FUNCTION_BLOCK "Sim: from Global"   // FB26, SCL
{ S7_Optimized_Access := 'TRUE' }
VERSION : 0.1
   VAR_INPUT
      stns : "Station: All Stations";
   END_VAR
   VAR_IN_OUT
      simStations : "Simulated Stations";
   END_VAR
   VAR
      old : Struct
         nextGrp : Bool;
         prevGrp : Bool;
      END_STRUCT;
   END_VAR
   VAR_TEMP
      animate : USInt;
      btnCount : Int;
      currentBtn : Bool;
      dzLabel : WString;
      firstStn : Int;
      i : Int;
      intBox : Int;
      j : Int;
      kp8Color : DWord;
      label : WString;
      oldBtn : Bool;
      pSim : Int;
      pStn : Int;
   END_VAR
   VAR CONSTANT
      space : WString := WSTRING#' ';
      lead0 : WString := WSTRING#'0';
      volvo16 : WString := WSTRING#'VOLVO 16';
   END_VAR
BEGIN
   REGION "COPY TO LOCAL"
       #firstStn := #simStations.firstStn;
   END_REGION

   REGION "RESOLVE STATION POINTER"

       REGION "PROCESS NEXT GROUP PRESS"

           REGION "COPY TO LOCAL"
               #currentBtn := #simStations.down.actuate;
               #oldBtn := #old.nextGrp;
           END_REGION

           REGION "FALLING EDGE OF NEXT GROUP"
               IF NOT #currentBtn AND #oldBtn THEN

                   REGION "INCREMENT FIRST STATION"
                       #firstStn += "simKP8Count";
                   END_REGION

                   REGION "UPPER LIMIT ROLL OVER"
                       IF #firstStn > "STATION_COUNT" THEN
                           #firstStn -= "STATION_COUNT" + 1;
                       END_IF;
                   END_REGION

               END_IF;
           END_REGION

           REGION "NEXT GROUP CHANGE DETECTION"
               #old.nextGrp := #currentBtn;
           END_REGION

       END_REGION

       REGION "PROCESS PREVIOUS GROUP PRESS"

           REGION "COPY TO LOCAL"
               #currentBtn := #simStations.up.actuate;
               #oldBtn := #old.prevGrp;
           END_REGION

           REGION "FALLING EDGE OF PREVIOUS GROUP"
               IF NOT #currentBtn AND #oldBtn THEN

                   REGION "DECREMENT FIRST STATION"
                       #firstStn -= "simKP8Count";
                   END_REGION

                   REGION "LOWER LIMIT ROLL OVER"
                       IF #firstStn < 0 THEN
                           #firstStn += "STATION_COUNT" + 1;
                       END_IF;
                   END_REGION

               END_IF;
           END_REGION

           REGION "PREVIOUS GROUP CHANGE DETECTION"
               #old.prevGrp := #currentBtn;
           END_REGION

       END_REGION

   END_REGION

   REGION "FOR EACH BUTTON"
       FOR #i := 0 TO 11 DO

           REGION "CALCULATE POINTER"
               #pStn := #i + #firstStn;
               #pSim := #i;
           END_REGION

           REGION "UPPER LIMIT ROLL OVER"
               IF #pStn > "STATION_COUNT" THEN
                   #pStn := #firstStn + #i - "STATION_COUNT" - 1;
               END_IF;
           END_REGION

           REGION "COPY TO LOCAL"
               #kp8Color := #stns.stn[#pStn].wipCmpts.ioData.kp8.tempOut;
           END_REGION

           REGION "LABEL STATIONS"

               REGION "DETERMINE LINE LABEL"
                   #label := #stns.stn[#pStn].id.lineName;
                   IF #label = #volvo16 THEN
                       #label := WSTRING#'V16';
                   END_IF;
               END_REGION

               REGION "DETERMINE DROP ZONE LABEL"
                   #intBox := USINT_TO_INT(#stns.stn[#pStn].id.dropZone);
                   IF #intBox <= 9 THEN
                       #dzLabel := CONCAT_WSTRING(IN1 := #lead0,
                                                  IN2 := "Strip Sign"(INT_TO_WSTRING(#intBox)));
                   END_IF;
                   IF #intBox >= 10 THEN
                       #dzLabel := "Strip Sign"(INT_TO_WSTRING(#intBox));
                   END_IF;
               END_REGION

               REGION "WRITE LABEL"
                   #label := CONCAT_WSTRING(IN1 := #label,
                                            IN2 := #space,
                                            IN3 := #dzLabel);
                   #simStations.me[#pSim].stn.label := #label;
               END_REGION

           END_REGION

           REGION "ANIMATE STATION LABEL"
               #simStations.me[#pSim].stn.animate := "GRAY_BACKGROUND";
           END_REGION

           REGION "FOR EACH BUTTON"
               FOR #j := 0 TO "BUTTON_COUNT" DO

                   REGION "COLOR BUTTONS"
                       #animate := "KP8 Driver: HMI Emulator: Animation"(kp8Color := #kp8Color,
                                                                btnNumber := #j);
                       #simStations.me[#pSim].btn.animate[#j] := #animate;
                   END_REGION

                   REGION "WRITE BUTTON LABELS"
                       #intBox := "Pointer Calc: KP8 Labels"(#j);
                       #label := "Strip Sign"(INT_TO_WSTRING(#intBox));
                       #simStations.me[#pSim].btn.labels[#j] := #label;
                   END_REGION

               END_FOR;
           END_REGION

       END_FOR;
   END_REGION

   REGION "SAVE FIRST STATION"
       #simStations.firstStn := #firstStn;
   END_REGION

   REGION "ANIMATE NEXT GROUP PRESS"
       #simStations.down.animate := "Bool.Animate"(true_color := "GREEN_LIGHT_BACKGROUND",
                                                   false_color := "GRAY_BACKGROUND",
                                                   evaluation_signal := #simStations.down.actuate);
   END_REGION

   REGION "ANIMATE PREV GROUP PARESS"
       #simStations.up.animate := "Bool.Animate"(true_color := "GREEN_LIGHT_BACKGROUND",
                                                 false_color := "GRAY_BACKGROUND",
                                                 evaluation_signal := #simStations.up.actuate);
   END_REGION
END_FUNCTION_BLOCK

FUNCTION "Sim: to Global" : Void   // FC23, SCL
{ S7_Optimized_Access := 'TRUE' }
VERSION : 0.1
   VAR_INPUT
      simStns : "Simulated Stations";
   END_VAR
   VAR_IN_OUT
      stations : "Station: All Stations";
   END_VAR
   VAR_TEMP
      i : Int;
      j : Int;
      pSim : Int;
      pStn : Int;
   END_VAR
BEGIN
   REGION "COPY TO LOCAL"
       // #btnCount := "btnCount";
       // #firstStn := #simStns.firstStn;
       // #simKP8Count := "simKP8Count";
       // #stnCount := "stnCount";
   END_REGION

   REGION "FOR EACH STATION"
       FOR #i := 0 TO "simKP8Count" DO

           REGION "CALCULATE POINTER"
               #pStn := #i + #simStns.firstStn;
               #pSim := #i;
           END_REGION

           REGION "UPPER LIMIT ROLL OVER"
               IF #pStn > "STATION_COUNT" THEN
                   #pStn := #simStns.firstStn + #i - "STATION_COUNT" - 1;
               END_IF;
           END_REGION

           REGION "COPY SIMULATED PRESSES"
               #stations.stn[#pStn].wipCmpts.ioData.kp8.input.%B1 := #simStns.me[#pSim].btn.actuate;
           END_REGION

       END_FOR;
   END_REGION
END_FUNCTION

FUNCTION "Sim: KP8 Animations" : Word   // FC84, SCL
{ S7_Optimized_Access := 'TRUE' }
VERSION : 0.1
   VAR_INPUT
      pbs : DWord;
   END_VAR
   VAR_TEMP
      ret : Word;
   END_VAR
BEGIN
   #"Sim: KP8 Animations".%B1 := #pbs.%B0;
   #"Sim: KP8 Animations".%B0 := #pbs.%B1;
END_FUNCTION

// folder: Flags

FUNCTION_BLOCK "Flag.New_PN_Code"   // FB3, SCL
{ S7_Optimized_Access := 'TRUE' }
VERSION : 0.1
   VAR_IN_OUT
      stns : "Station: All Stations";
   END_VAR
   VAR
      old : Struct
         pnCode : Array[0.."STATION_COUNT"] of Struct
            me : Array[0.."BUTTON_COUNT"] of DInt;
         END_STRUCT;
      END_STRUCT;
   END_VAR
   VAR_TEMP
      pStn : Int;
      ret : Bool;
   END_VAR
BEGIN
   REGION "FOR EACH STATION"
       FOR #pStn := 0 TO "STATION_COUNT" DO

           REGION "ON PART NUMBER CHANGE"
               IF #stns.stn[#pStn].wipCmpts.pnCode <> #old.pnCode[#pStn].me THEN

                   REGION "SET FLAG"
                       #ret := TRUE;
                   END_REGION

               END_IF;
           END_REGION

           REGION "SAVE FLAG"
               #stns.stn[#pStn].wipCmpts.flags.newPN := #ret;
           END_REGION

           REGION "CHANGE DETECTION"
               #old.pnCode[#pStn].me := #stns.stn[#pStn].wipCmpts.pnCode;
           END_REGION

       END_FOR;
   END_REGION
END_FUNCTION_BLOCK

FUNCTION_BLOCK "Flag.State_Transition"   // FB4, SCL
{ S7_Optimized_Access := 'TRUE' }
VERSION : 0.1
   VAR_IN_OUT
      stns : "Station: All Stations";
   END_VAR
   VAR
      old : Struct
         stn : Array[0.."STATION_COUNT"] of Struct
            orderState : Array[0.."BUTTON_COUNT"] of Int;
         END_STRUCT;
      END_STRUCT;
   END_VAR
   VAR_TEMP
      pStn : Int;
      pBtn : Int;
      ret : Bool;
   END_VAR
BEGIN
   REGION "FOR EACH STATION"
       FOR #pStn := 0 TO "STATION_COUNT" DO

           REGION "IGNORE WIP LOAD CYCLE"
               IF NOT #stns.stn[#pStn].flags.wipSwapped THEN

                   REGION "FOR EACH BUTTON"
                       FOR #pBtn := 0 TO "BUTTON_COUNT" DO

                           REGION "RESET RETURN"
                               #ret := FALSE;
                           END_REGION

                           REGION "ON CHANGE IN STATE"
                               IF #stns.stn[#pStn].wipCmpts.orderState[#pBtn] <> #old.stn[#pStn].orderState[#pBtn] THEN

                                   REGION "SET STATE TRANSITION FLAG"
                                       #ret := true;
                                   END_REGION

                               END_IF;
                           END_REGION

                           REGION "SAVE FLAG"
                               #stns.stn[#pStn].flags.stateTransition[#pBtn] := #ret;
                           END_REGION

                       END_FOR;
                   END_REGION

               END_IF;
           END_REGION

           REGION "CHANGE DETECTION"
               #old.stn[#pStn].orderState := #stns.stn[#pStn].wipCmpts.orderState;
           END_REGION

       END_FOR;
   END_REGION
END_FUNCTION_BLOCK

FUNCTION_BLOCK "Flag"   // FB5, SCL
{ S7_Optimized_Access := 'TRUE' }
VERSION : 0.1
   VAR_INPUT
      pnLib : "Recipe: PN Text Library";
      screen_number : Int;
   END_VAR
   VAR_IN_OUT
      stns : "Station: All Stations";
      savedStns : "Recipe: HMI Stations Saved Wips";
   END_VAR
   VAR
      _i : Int;
      "inst New PN Code" : "Flag.New_PN_Code";
      "inst Flag: State Transition" : "Flag.State_Transition";
      "inst Flag: Wip Deselect" : "Flag.Wip_Deselect";
      "inst Flag: Wip Swapped" : "Flag.Wip_Swapped";
   END_VAR
BEGIN
   REGION "NEW PART NUMBER ASSIGNED"
       #"inst New PN Code"(#stns);
   END_REGION

   REGION "PART NUMBER VALIDATION"
       "Flag.PN_Good"(pnLib := #pnLib,
                       stns := #stns);
   END_REGION

   REGION "WIP SWAPPED"
       #"inst Flag: Wip Swapped"(#stns);
   END_REGION

   REGION "STATE TRANSITIONS"
       #"inst Flag: State Transition"(#stns);
   END_REGION

   REGION "WIP DESELECTION"
       #"inst Flag: Wip Deselect"(#savedStns);
   END_REGION

   REGION "IN SETTINGS SCREEN"
       FOR #_i := 0 TO "STATION_COUNT" DO
           #stns.stn[#_i].wipCmpts.flags.inSettingsScreen := "Flag.In_Settings_Screen"(#screen_number);
       END_FOR;
   END_REGION
END_FUNCTION_BLOCK

FUNCTION_BLOCK "Flag.Wip_Swapped"   // FB10, SCL
{ S7_Optimized_Access := 'TRUE' }
VERSION : 0.1
   VAR_IN_OUT
      stns : "Station: All Stations";
   END_VAR
   VAR
      old : Struct
         wipIndex : Array[0.."STATION_COUNT"] of DInt;
      END_STRUCT;
   END_VAR
   VAR_TEMP
      pStn : Int;
      ret : Bool;
   END_VAR
BEGIN
   REGION "FOR EACH STATION"
       FOR #pStn := 0 TO "STATION_COUNT" DO

           REGION "ON WIP CHANGE"
               IF #stns.stn[#pStn].wipData.index <> #old.wipIndex[#pStn] THEN

                   REGION "SET FLAG"
                       #ret := TRUE;
                   END_REGION

                   REGION "SAVE FLAG"
                       #stns.stn[#pStn].wipCmpts.flags.newPN := #ret;
                   END_REGION

               END_IF;
           END_REGION

           REGION "CHANGE DETECTION"
               #old.wipIndex[#pStn] := #stns.stn[#pStn].wipData.index;
           END_REGION

       END_FOR;
   END_REGION
END_FUNCTION_BLOCK

FUNCTION_BLOCK "Flag.Wip_Deselect.Flag Pulse"   // FB17, SCL
{ S7_Optimized_Access := 'TRUE' }
VERSION : 0.1
   VAR_INPUT
      remaining : Real;
      reset : Bool;
   END_VAR
   VAR_IN_OUT
      flag : Bool;
   END_VAR
   VAR RETAIN
      hasBeenFlipped : Bool;
   END_VAR
BEGIN
   #flag := FALSE;

   IF #reset THEN
       #hasBeenFlipped := FALSE;
       RETURN;
   END_IF;

   IF #remaining >= 0.0 THEN
       #hasBeenFlipped := FALSE;
       RETURN;
   END_IF;

   IF NOT #hasBeenFlipped THEN
       IF #remaining < 0.0 THEN
           #hasBeenFlipped := TRUE;
           #flag := TRUE;
       END_IF;
   END_IF;
END_FUNCTION_BLOCK

FUNCTION_BLOCK "Flag.Wip_Deselect"   // FB18, SCL
{ S7_Optimized_Access := 'TRUE' }
VERSION : 0.1
   VAR_IN_OUT
      savedStns : "Recipe: HMI Stations Saved Wips";
   END_VAR
   VAR
      "inst Flag Pulses" : Array[0.."STATION_COUNT", 0.."WIP_COUNT"] of "Flag.Wip_Deselect.Flag Pulse";
   END_VAR
   VAR_TEMP
      pStn : Int;
      pWip : Int;
   END_VAR
BEGIN
   REGION "FOR EACH STATION"
       FOR #pStn := 0 TO "HMI_STATION_COUNT" DO

           REGION "FOR EACH WIP"
               FOR #pWip := 0 TO "WIP_COUNT" DO

                   REGION "FLAG PULSE"
                       #"inst Flag Pulses"[#pStn, #pWip](remaining := #savedStns.stn[#pStn].wip[#pWip].timers.wdsRemaining,
                                                         flag := #savedStns.stn[#pStn].wip[#pWip].flags.clearWipRequest);
                   END_REGION

               END_FOR;
           END_REGION

       END_FOR;
   END_REGION
END_FUNCTION_BLOCK

FUNCTION "Flag.PN_Good" : Void   // FC13, SCL
{ S7_Optimized_Access := 'TRUE' }
VERSION : 0.1
   VAR_INPUT
      pnLib : "Recipe: PN Text Library";
   END_VAR
   VAR_IN_OUT
      stns : "Station: All Stations";
   END_VAR
   VAR_TEMP
      pStn : Int;
      pBtn : Int;
      pnGood : Bool;
   END_VAR
BEGIN
   REGION "FOR EACH STATION"
       FOR #pStn := 0 TO "STATION_COUNT" DO

           REGION "FOR EACH BUTTON"
               FOR #pBtn := 0 TO "BUTTON_COUNT" DO

                   REGION "ON NEW PN"
                       IF #stns.stn[#pStn].wipCmpts.flags.newPN THEN

                           REGION "VALIDATE PN"
                               #pnGood := "Validate PN"(pnCode := #stns.stn[#pStn].wipCmpts.pnCode[#pBtn],
                                                        pnLib := #pnLib);
                           END_REGION

                           REGION "SAVE TO FLAG"
                               #stns.stn[#pStn].wipCmpts.flags.pnGood[#pBtn] := #pnGood;
                           END_REGION

                       END_IF;
                   END_REGION

               END_FOR;
           END_REGION

       END_FOR;
   END_REGION
END_FUNCTION

FUNCTION "Flag.In_Settings_Screen" : Bool   // FC294, SCL
{ S7_Optimized_Access := 'TRUE' }
VERSION : 0.1
   VAR_INPUT
      screen_number : Int;
   END_VAR
   VAR CONSTANT
      SETTINGS_SCREEN_NUMBER : Int := 2;
   END_VAR
BEGIN
   #"Flag.In_Settings_Screen" := #screen_number = #SETTINGS_SCREEN_NUMBER;
END_FUNCTION

// folder: From Excel

FUNCTION_BLOCK "From Excel"   // FB8, SCL
{ S7_Optimized_Access := 'TRUE' }
VERSION : 0.1
   VAR_INPUT
      codeLib : "From Excel: Data";
   END_VAR
   VAR_IN_OUT
      stns : "Station: All Stations";
      svdHMIStnWips : "Recipe: HMI Stations Saved Wips";
   END_VAR
   VAR
      operation_complete : Bool;
      start : Bool;
      states : "Initialize Excel Data: States";
   END_VAR
BEGIN
   REGION "STATE MACHINE"
       "Initialize Excel Data: State Machine"(start := "FirstScan" OR #start,
                                              states := #states,
                                              operation_complete := #operation_complete);
   END_REGION

   REGION "LOAD PART NUMBER CODES TO KP8 STATIONS"
       IF #states.pn_code_to_kp8_station THEN
           "From Excel: PN Code to KP8 Stations"(code_library := #codeLib,
                                                 stations := #stns,
                                                 operation_complete := #operation_complete);
       END_IF;
   END_REGION

   REGION "LOAD PART NUMBER CODES TO SAVED WIPS"
       IF #states.pn_code_to_saved_wips THEN
           "From Excel: PN Code to HMI Station Saved Wips"(code_libarary := #codeLib,
                                                           saved_wip_stations := #svdHMIStnWips,
                                                           operation_complete := #operation_complete);
       END_IF;
   END_REGION

   REGION "LOAD WIP CODES TO SAVED WIPS"
       IF #states.wip_code_to_saved_wips THEN
           "From Excel: Wip Code to HMI Station Saved WIps"(excel_code_library := #codeLib,
                                                            saved_wip_stations := #svdHMIStnWips,
                                                            operation_complete := #operation_complete);
       END_IF;
   END_REGION

   REGION "LOAD ACTIVE WIP TO HMI STATION LIST"
       IF #states.active_wip_to_hmi_station_list THEN
           "From Excel: HMI Stations Load Active WIP"(excel_code_library := #codeLib,
                                                      stations := #stns,
                                                      operation_complete := #operation_complete);
       END_IF;
   END_REGION

   REGION "LOAD ACTIVE WIP TO MASTER STATION LIST"
       IF #states.active_wip_to_master_station_list THEN
           "HMI Station: Load Active WIP into Master Station List"(operation_complete := #operation_complete);
       END_IF;
   END_REGION
END_FUNCTION_BLOCK

FUNCTION "From Excel: PN Code to KP8 Stations" : Void   // FC58, SCL
{ S7_Optimized_Access := 'TRUE' }
VERSION : 0.1
   VAR_INPUT
      code_library : "From Excel: Data";
   END_VAR
   VAR_IN_OUT
      stations : "Station: All Stations";
      operation_complete : Bool;
   END_VAR
   VAR_TEMP
      pointer_source : Int;
      pointer_destination : Int;
   END_VAR
BEGIN
   REGION "KP8 STATIONS
       FOR #pointer_source := 0 TO UDINT_TO_INT("Array.Any.Length"(#code_library.kp8Stns) - 1) DO
           #pointer_destination := #code_library.kp8Stns[#pointer_source].pStn;
           IF #pointer_destination = -1 THEN
               EXIT;
           END_IF;
           #stations.stn[#pointer_destination].wipCmpts.pnCode := #code_library.kp8Stns[#pointer_source].pnCode;
       END_FOR;
       #operation_complete := TRUE;
   END_REGION
END_FUNCTION

FUNCTION "From Excel: PN Code to HMI Station Saved Wips" : Void   // FC61, SCL
{ S7_Optimized_Access := 'TRUE' }
VERSION : 0.1
   VAR_INPUT
      code_libarary : "From Excel: Data";
   END_VAR
   VAR_IN_OUT
      saved_wip_stations : "Recipe: HMI Stations Saved Wips";
      operation_complete : Bool;
   END_VAR
   VAR_TEMP
      pointer_source_station : Int;
      pointer_destination_station : Int;
      pointer_wip : Int;
   END_VAR
BEGIN
   REGION "HMI STATIONS"
       FOR #pointer_source_station := 0 TO UDINT_TO_INT("Array.Any.Length"(#code_libarary.hmiStns) - 1) DO
           #pointer_destination_station := #code_libarary.hmiStns[#pointer_source_station].pStn;
           IF #pointer_destination_station = -1 THEN
               EXIT;
           END_IF;
           FOR #pointer_wip := 0 TO "WIP_COUNT" DO
               #saved_wip_stations.stn[#pointer_source_station].wip[#pointer_wip].pnCode :=
                   #code_libarary.hmiStns[#pointer_source_station].wip[#pointer_wip].pnCode;
           END_FOR;
       END_FOR;
       #operation_complete := TRUE;
   END_REGION
END_FUNCTION

FUNCTION "From Excel: HMI Stations Load Active WIP" : Void   // FC62, SCL
{ S7_Optimized_Access := 'TRUE' }
VERSION : 0.1
   VAR_INPUT
      excel_code_library : "From Excel: Data";
   END_VAR
   VAR_IN_OUT
      stations : "Station: All Stations";
      operation_complete : Bool;
   END_VAR
   VAR_TEMP
      pointer_source : Int;
      pointer_destination : Int;
   END_VAR
BEGIN
   REGION "HMI STATIONS"
       FOR #pointer_source := 0 TO UDINT_TO_INT("Array.Any.Length"(#excel_code_library.hmiStns) - 1) DO
           #pointer_destination := #excel_code_library.hmiStns[#pointer_source].pStn;
           IF #pointer_destination = -1 THEN
               EXIT;
           END_IF;
           #stations.stn[#pointer_destination].wipCmpts.pnCode := #excel_code_library.hmiStns[#pointer_source].wip[0].pnCode;
       END_FOR;
       #operation_complete := TRUE;
   END_REGION
END_FUNCTION

FUNCTION "From Excel: Wip Code to HMI Station Saved WIps" : Void   // FC63, SCL
{ S7_Optimized_Access := 'TRUE' }
VERSION : 0.1
   VAR_INPUT
      excel_code_library : "From Excel: Data";
   END_VAR
   VAR_IN_OUT
      saved_wip_stations : "Recipe: HMI Stations Saved Wips";
      operation_complete : Bool;
   END_VAR
   VAR_TEMP
      "pointer_source _station" : Int;
      pointer_destination_station : Int;
      pointer_wip : Int;
   END_VAR
BEGIN
   REGION "HMI STATIONS"
       FOR #"pointer_source _station" := 0 TO UDINT_TO_INT("Array.Any.Length"(#excel_code_library.hmiStns) - 1) DO
           FOR #pointer_wip := 0 TO "WIP_COUNT" DO
               #saved_wip_stations.stn[#"pointer_source _station"].wip[#pointer_wip].wip.code :=
                   #excel_code_library.hmiStns[#"pointer_source _station"].wip[#pointer_wip].wipCode;
           END_FOR;
       END_FOR;
       #operation_complete := TRUE;
   END_REGION
END_FUNCTION

FUNCTION "Initialize Excel Data: State Machine" : Void   // FC148, SCL
{ S7_Optimized_Access := 'TRUE' }
VERSION : 0.1
   VAR_INPUT
      start : Bool;
   END_VAR
   VAR_IN_OUT
      states : "Initialize Excel Data: States";
      operation_complete : Bool;
   END_VAR
   VAR_TEMP
      clear_states : "Initialize Excel Data: States";
   END_VAR
BEGIN
   REGION "LOAD PART NUMBER CODES TO KP8 STATIONS"
       IF #start AND NOT #operation_complete AND "Initialize Excel Data: All States False"(#states) THEN
           #states := #clear_states;
           #states.pn_code_to_kp8_station := TRUE;
           #operation_complete := FALSE;
       END_IF;
   END_REGION

   REGION "LOAD PART NUMBER CODES TO SAVED WIPS"
       IF #states.pn_code_to_kp8_station AND #operation_complete THEN
           #states := #clear_states;
           #states.pn_code_to_saved_wips := TRUE;
           #operation_complete := FALSE;
       END_IF;
   END_REGION

   REGION "LOAD WIP CODES TO SAVED WIPS"
       IF #states.pn_code_to_saved_wips AND #operation_complete THEN
           #states := #clear_states;
           #states.wip_code_to_saved_wips := TRUE;
           #operation_complete := FALSE;
       END_IF;
   END_REGION

   REGION "LOAD ACTIVE WIP TO HMI STATION LIST"
       IF #states.wip_code_to_saved_wips AND #operation_complete THEN
           #states := #clear_states;
           #states.active_wip_to_hmi_station_list := TRUE;
           #operation_complete := FALSE;
       END_IF;
   END_REGION

   REGION "LOAD ACTIVE WIP TO MASTER STATION LIST"
       IF #states.active_wip_to_hmi_station_list AND #operation_complete THEN
           #states := #clear_states;
           #states.active_wip_to_master_station_list := TRUE;
           #operation_complete := FALSE;
       END_IF;
   END_REGION

   REGION "COMPLETE"
       IF #states.active_wip_to_master_station_list AND #operation_complete THEN
           #states := #clear_states;
           #operation_complete := FALSE;
       END_IF;
   END_REGION
END_FUNCTION

FUNCTION "Initialize Excel Data: All States False" : Bool   // FC149, SCL
{ S7_Optimized_Access := 'TRUE' }
VERSION : 0.1
   VAR_INPUT
      states : "Initialize Excel Data: States";
   END_VAR
   VAR_TEMP
      ret : Bool;
   END_VAR
BEGIN
   IF NOT #states.active_wip_to_hmi_station_list AND
       NOT #states.pn_code_to_kp8_station AND
       NOT #states.active_wip_to_master_station_list AND
       NOT #states.pn_code_to_saved_wips AND
       NOT #states.wip_code_to_saved_wips THEN
       #ret := TRUE;
   END_IF;
   #"Initialize Excel Data: All States False" := #ret;
END_FUNCTION

// folder: Global/Physical

FUNCTION "Physical to Global" : Void   // FC1, LAD
{ S7_Optimized_Access := 'TRUE' }
VERSION : 0.1
   VAR_IN_OUT
      stations : "Station: All Stations";
   END_VAR
   VAR_TEMP
      i : Int;
      kp8In : DWord;
   END_VAR
BEGIN

REGION Network 1 (SCL): MAIN LOOP
   FOR #i := 0 TO "STATION_COUNT" DO

       CASE #i OF
           "VOLVO 16 01":
               #kp8In := "VOLVO 16 01 KP8 In";
           "VOLVO 16 02":
               #kp8In := "VOLVO 16 02 KP8 In";
           "VOLVO 16 03":
               #kp8In := "VOLVO 16 03 KP8 In";
           "VOLVO 16 04":
               #kp8In := "VOLVO 16 04 KP8 In";
           "VOLVO 16 05":
               #kp8In := "VOLVO 16 05 KP8 In";
           "VOLVO 16 06":
               #kp8In := "VOLVO 16 06 KP8 In";
           "VOLVO 16 07":
               #kp8In := "VOLVO 16 07 KP8 In";
           "VOLVO 16 08":
               #kp8In := "VOLVO 16 08 KP8 In";
           "VOLVO 16 09":
               #kp8In := "VOLVO 16 09 KP8 In";
           "VOLVO 16 10":
               #kp8In := "VOLVO 16 10 KP8 In";
           "VOLVO 16 11":
               #kp8In := "VOLVO 16 11 KP8 In";
           "CHM 01":
               #kp8In := "CHM 01 KP8 In";
           "CHM 02":
               #kp8In := "CHM 02 KP8 In";
           "CHM 03":
               #kp8In := "CHM 03 KP8 In";
           "CHM 04":
               #kp8In := "CHM 04 KP8 In";
           "CHM 05":
               #kp8In := "CHM 05 KP8 In";
           "CDO 01":
               #kp8In := "CDO 01 KP8 In";
           "CDO 02":
               #kp8In := "CDO 02 KP8 In";
           "CDO 03":
               #kp8In := "CDO 03 KP8 In";
           "BFL 01":
               #kp8In := "BFL 01 KP8 In";
           "BFL 02":
               #kp8In := "BFL 02 KP8 In";
           "BFL 03":
               #kp8In := "BFL 03 KP8 In";
           "LGS 01":
               #kp8In := "LGS 01 KP8 In";
           "LGS 02":
               #kp8In := "LGS 02 KP8 In";
           "LGS 03":
               #kp8In := "LGS 03 KP8 In";
           "CV 01":
               #kp8In := "CV 01 KP8 In";
           "CV 02":
               #kp8In := "CV 02 KP8 In";
           "CV 03":
               #kp8In := "CV 03 KP8 In";
           "CV 04":
               #kp8In := "CV 04 KP8 In";
           "PC 01":
               #kp8In := "PC 01 KP8 In"; 
           "PC 02":
               #kp8In := "PC 02 KP8 In";
       END_CASE;

       #stations.stn[#i].wipCmpts.ioData.kp8.input := #kp8In.%W1;

   END_FOR;
END_REGION
END_FUNCTION

FUNCTION "Global to Physical" : Void   // FC5, LAD
{ S7_Optimized_Access := 'TRUE' }
VERSION : 0.1
   VAR_IN_OUT
      stations : "Station: All Stations";
   END_VAR
   VAR_TEMP
      i : Int;
      j : Int;
      ET200SP : DWord;
      "KP8 In" : DWord;
      "KP8 Out" : DWord;
      Card : Int;
      stnCount : Int;
   END_VAR
BEGIN

REGION Network 1 (SCL): MAIN LOOP
   FOR #i := 0 TO "STATION_COUNT" DO

       #ET200SP := #stations.stn[#i].wipCmpts.ioData.stkLight;
       #"KP8 Out" := #stations.stn[#i].wipCmpts.ioData.kp8.tempOut;

       CASE #i OF
           "VOLVO 16 01":
               "VOLVO 16 01 IO" := #ET200SP;
               "VOLVO 16 01 KP8 Out" := #"KP8 Out";
           "VOLVO 16 02":
               "VOLVO 16 02 IO" := #ET200SP;
               "VOLVO 16 02 KP8 Out" := #"KP8 Out";
           "VOLVO 16 03":
               "VOLVO 16 03 IO" := #ET200SP;
               "VOLVO 16 03 KP8 Out" := #"KP8 Out";
           "VOLVO 16 04":
               "VOLVO 16 04 IO" := #ET200SP;
               "VOLVO 16 04 KP8 Out" := #"KP8 Out";
           "VOLVO 16 05":
               "VOLVO 16 05 IO" := #ET200SP;
               "VOLVO 16 05 KP8 Out" := #"KP8 Out";
           "VOLVO 16 06":
               "VOLVO 16 06 IO" := #ET200SP;
               "VOLVO 16 06 KP8 Out" := #"KP8 Out";
           "VOLVO 16 07":
               "VOLVO 16 07 IO" := #ET200SP;
               "VOLVO 16 07 KP8 Out" := #"KP8 Out";
           "VOLVO 16 08":
               "VOLVO 16 08 IO" := #ET200SP;
               "VOLVO 16 08 KP8 Out" := #"KP8 Out";
           "VOLVO 16 09":
               "VOLVO 16 09 IO" := #ET200SP;
               "VOLVO 16 09 KP8 Out" := #"KP8 Out";
           "VOLVO 16 10":
               "VOLVO 16 10 IO" := #ET200SP;
               "VOLVO 16 10 KP8 Out" := #"KP8 Out";
           "VOLVO 16 11":
               "VOLVO 16 11 IO" := #ET200SP;
               "VOLVO 16 11 KP8 Out" := #"KP8 Out";
           "CHM 01":
               "CHM 01 IO" := #ET200SP;
               "CHM 01 KP8 Out" := #"KP8 Out";
           "CHM 02":
               "CHM 02 IO" := #ET200SP;
               "CHM 02 KP8 Out" := #"KP8 Out";
           "CHM 03":
               "CHM 03 IO" := #ET200SP;
               "CHM 03 KP8 Out" := #"KP8 Out";
           "CHM 04":
               "CHM 04 IO" := #ET200SP;
               "CHM 04 KP8 Out" := #"KP8 Out";
           "CHM 05":
               "CHM 05 IO" := #ET200SP;
               "CHM 05 KP8 Out" := #"KP8 Out";
           "CDO 01":
               "CDO 01 IO" := #ET200SP;
               "CDO 01 KP8 Out" := #"KP8 Out";
           "CDO 02":
               "CDO 02 IO" := #ET200SP;
               "CDO 02 KP8 Out" := #"KP8 Out";
           "CDO 03":
               "CDO 03 IO" := #ET200SP;
               "CDO 03 KP8 Out" := #"KP8 Out";
           "BFL 01":
               "BFL 01 IO" := #ET200SP;
               "BFL 01 KP8 Out" := #"KP8 Out";
           "BFL 02":
               "BFL 02 IO" := #ET200SP;
               "BFL 02 KP8 Out" := #"KP8 Out";
           "BFL 03":
               "BFL 03 IO" := #ET200SP;
               "BFL 03 KP8 Out" := #"KP8 Out";
           "LGS 01":
               "LGS 01 IO" := #ET200SP;
               "LGS 01 KP8 Out" := #"KP8 Out";
           "LGS 02":
               "LGS 02 IO" := #ET200SP;
               "LGS 02 KP8 Out" := #"KP8 Out";
           "LGS 03":
               "LGS 03 IO" := #ET200SP;
               "LGS 03 KP8 Out" := #"KP8 Out";
           "CV 01":
               "CV 01 IO" := #ET200SP;
               "CV 01 KP8 Out" := #"KP8 Out";
           "CV 02":
               "CV 02 IO" := #ET200SP;
               "CV 02 KP8 Out" := #"KP8 Out";
           "CV 03":
               "CV 03 IO" := #ET200SP;
               "CV 03 KP8 Out" := #"KP8 Out";
           "CV 04":
               "CV 04 IO" := #ET200SP;
               "CV 04 KP8 Out" := #"KP8 Out";
           "PC 01":
               "PC 01 IO" := #ET200SP;
               "PC 01 KP8 Out" := #"KP8 Out";
           "PC 02":
               "PC 02 IO" := #ET200SP;
               "PC 02 KP8 Out" := #"KP8 Out";

       END_CASE;

   END_FOR;
END_REGION
END_FUNCTION

// folder: Linked List

FUNCTION_BLOCK "Linked List"   // FB29, SCL
{ S7_Optimized_Access := 'TRUE' }
VERSION : 0.1
   VAR_IN_OUT
      interface : "Linked List: Method Interface";
   END_VAR
   VAR
      list : "Linked List: List";
   END_VAR
   VAR CONSTANT
      TERMINAL_BEHAVIOR : String := 'open';
   END_VAR
BEGIN
   REGION "APPEND"
       IF #interface.append.in.request THEN
           "Linked List: Append"(terminal_behavior := #TERMINAL_BEHAVIOR,
                                 commands := #interface.append,
                                 list := #list);
       END_IF;
   END_REGION

   REGION "DELETE"
       IF #interface.delete.in.request THEN
           "Linked List: Delete"(commands := #interface.delete,
                                 list := #list);
       END_IF;
   END_REGION

   REGION "DISPLAY"
       IF #interface.display.in.request THEN
           "Linked List: Display"(commands := #interface.display,
                                  list := #list);
       END_IF;
   END_REGION

   REGION "INSERT"
       IF #interface.insert.in.request THEN
           "Linked List: Insert"(terminal_behavior := #TERMINAL_BEHAVIOR,
                                 commands := #interface.insert,
                                 list := #list);
       END_IF;
   END_REGION

   REGION "RESET"
       IF #interface.reset.in.request THEN
           "Linked List: Reset"(commands := #interface.reset,
                                list := #list);
       END_IF;
   END_REGION

   REGION "REVERSE"
       IF #interface.reverse.in.request THEN
           "Linked List: Reverse"(commands := #interface.reverse,
                                  list := #list);
       END_IF;
   END_REGION

   REGION "SEARCH"
       IF #interface.search.in.request THEN
           "Linked List: Search"(commands := #interface.search,
                                 list := #list);
       END_IF;
   END_REGION
END_FUNCTION_BLOCK

FUNCTION "Linked List: Private: Clear Node" : Void   // FC156, SCL
{ S7_Optimized_Access := 'TRUE' }
VERSION : 0.1
   VAR_IN_OUT
      node : "Linked List: Node";
   END_VAR
   VAR_TEMP
      ret : "Linked List: Node";
   END_VAR
BEGIN
   #ret.meta.key := "NULL_TOKEN";
   #ret.meta.next := "NULL_TOKEN";
   #node := #ret;
END_FUNCTION

FUNCTION "Linked List: Private: Get Head" : "Linked List: Node"   // FC157, SCL
{ S7_Optimized_Access := 'TRUE' }
VERSION : 0.1
   VAR_INPUT
      list : "Linked List: List";
   END_VAR
   VAR_TEMP
      pointer_list : DInt;
      ret : "Linked List: Node";
   END_VAR
BEGIN
   FOR #pointer_list := 0 TO "LINKED_LIST_LENGTH" DO
       IF #list.me[#pointer_list].meta.is_head THEN
           #ret := #list.me[#pointer_list];
           EXIT;
       END_IF;
   END_FOR;
   #"Linked List: Private: Get Head" := #ret;
END_FUNCTION

FUNCTION "Linked List: Private: Before" : Void   // FC158, SCL
{ S7_Optimized_Access := 'TRUE' }
VERSION : 0.1
   VAR_IN_OUT
      next_node : "Linked List: Node";   // next_node goes after node
      node : "Linked List: Node";   // node goes before next_node
   END_VAR
BEGIN
   #node.meta.next := #next_node.meta.key;
   IF #next_node.meta.is_head THEN
       #next_node.meta.is_head := FALSE;
       #node.meta.is_head := TRUE;
   END_IF;
END_FUNCTION

FUNCTION "Linked List: Private: Tail Swap" : Void   // FC159, SCL
{ S7_Optimized_Access := 'TRUE' }
VERSION : 0.1
   VAR_IN_OUT
      new_tail : "Linked List: Node";
      old_tail : "Linked List: Node";
   END_VAR
BEGIN
   #new_tail.meta.is_tail := TRUE;
   #old_tail.meta.is_tail := FALSE;
END_FUNCTION

FUNCTION "Linked List: Private: Head Swap" : Void   // FC160, SCL
{ S7_Optimized_Access := 'TRUE' }
VERSION : 0.1
   VAR_IN_OUT
      new_head : "Linked List: Node";
      old_head : "Linked List: Node";
   END_VAR
BEGIN
   #new_head.meta.is_head := TRUE;
   #old_head.meta.is_head := FALSE;
END_FUNCTION

FUNCTION "Linked List: Private: Get Next" : "Linked List: Node"   // FC161, SCL
{ S7_Optimized_Access := 'TRUE' }
VERSION : 0.1
   VAR_INPUT
      current : "Linked List: Node";
      list : "Linked List: List";
   END_VAR
   VAR_TEMP
      ret : "Linked List: Node";
   END_VAR
BEGIN
   "Linked List: Private: Clear Node"(#ret);
   IF #list.me[#current.meta.key].meta.next <> "NULL_TOKEN" THEN
       #ret := #list.me[#current.meta.next];
   END_IF;
   #"Linked List: Private: Get Next" := #ret;
END_FUNCTION

FUNCTION "Linked List: Private: Get Previous" : "Linked List: Node"   // FC162, SCL
{ S7_Optimized_Access := 'TRUE' }
VERSION : 0.1
   VAR_INPUT
      current : "Linked List: Node";
      list : "Linked List: List";
   END_VAR
   VAR_TEMP
      list_pointer : DInt;
      ret : "Linked List: Node";
   END_VAR
BEGIN
   "Linked List: Private: Clear Node"(#ret);
   FOR #list_pointer := 0 TO "LINKED_LIST_LENGTH" DO
       IF #list.me[#list_pointer].meta.next = #current.meta.key THEN
           #ret := #list.me[#list_pointer];
           EXIT;
       END_IF;
   END_FOR;
   #"Linked List: Private: Get Previous" := #ret;
END_FUNCTION

FUNCTION "Linked List: Private: After" : Void   // FC163, SCL
{ S7_Optimized_Access := 'TRUE' }
VERSION : 0.1
   VAR_IN_OUT
      node : "Linked List: Node";
      previous_node : "Linked List: Node";
   END_VAR
BEGIN
   #node.meta.next := #previous_node.meta.next;
   #previous_node.meta.next := #node.meta.key;
   IF #previous_node.meta.is_tail THEN
       #previous_node.meta.is_tail := FALSE;
       #node.meta.is_tail := TRUE;
   END_IF;
END_FUNCTION

FUNCTION "Linked List: Private: Head an Empty List" : Void   // FC164, SCL
{ S7_Optimized_Access := 'TRUE' }
VERSION : 0.1
   VAR_INPUT
      data : "Linked List: Node: Data";
      terminal_behavior : String;   // 'open': head's previous and tail's next are null nodes; 'closed': head's previous is tail, tail's next is head
   END_VAR
   VAR_IN_OUT
      list : "Linked List: List";
   END_VAR
BEGIN
   #list.me[0].data := #data;
   #list.me[0].meta.key := 0;
   IF #terminal_behavior = 'open' THEN
       #list.me[0].meta.next := "NULL_TOKEN";
   END_IF;
   IF #terminal_behavior = 'closed' THEN
       #list.me[0].meta.next := 0;
   END_IF;
   #list.me[0].meta.is_head := TRUE;
   #list.me[0].meta.is_tail := TRUE;
END_FUNCTION

FUNCTION "Linked List: Private: Is Empty" : Bool   // FC165, SCL
{ S7_Optimized_Access := 'TRUE' }
VERSION : 0.1
   VAR_INPUT
      list : "Linked List: List";
   END_VAR
   VAR_TEMP
      pointer_list : DInt;
      ret : Bool;
   END_VAR
BEGIN
   #ret := TRUE;
   FOR #pointer_list := 0 TO "LINKED_LIST_LENGTH" DO
       IF #list.me[#pointer_list].meta.key <> "NULL_TOKEN" THEN
           #ret := FALSE;
           EXIT;
       END_IF;
   END_FOR;
   #"Linked List: Private: Is Empty" := #ret;
END_FUNCTION

FUNCTION "Linked List: Private: Get Tail" : "Linked List: Node"   // FC166, SCL
{ S7_Optimized_Access := 'TRUE' }
VERSION : 0.1
   VAR_IN_OUT
      list : "Linked List: List";
   END_VAR
   VAR_TEMP
      pointer_list : Int;
      next_node : UInt;
      ret : "Linked List: Node";
   END_VAR
BEGIN
   FOR #pointer_list := 0 TO "LINKED_LIST_LENGTH" DO
       IF #list.me[#pointer_list].meta.is_tail THEN
           #ret := #list.me[#pointer_list];
           EXIT;
       END_IF;
   END_FOR;
   #"Linked List: Private: Get Tail" := #ret;
END_FUNCTION

FUNCTION "Linked List: Private: Is Full" : Bool   // FC167, SCL
{ S7_Optimized_Access := 'TRUE' }
VERSION : 0.1
   VAR_INPUT
      list : "Linked List: List";
   END_VAR
   VAR_TEMP
      pointer_list : DInt;
      ret : Bool;
   END_VAR
BEGIN
   #ret := TRUE;
   FOR #pointer_list := 0 TO "LINKED_LIST_LENGTH" DO
       IF #list.me[#pointer_list].meta.key = "NULL_TOKEN" THEN
           #ret := FALSE;
           EXIT;
       END_IF;
   END_FOR;
   #"Linked List: Private: Is Full" := #ret;
END_FUNCTION

FUNCTION "Linked List: Private: Next Empty Node" : DInt   // FC168, SCL
{ S7_Optimized_Access := 'TRUE' }
VERSION : 0.1
   VAR_IN_OUT
      list : "Linked List: List";
   END_VAR
   VAR_TEMP
      node : "Linked List: Node";
      pointer_list : Int;
      ret : DInt;
   END_VAR
BEGIN
   #ret := "NULL_TOKEN";
   FOR #pointer_list := 0 TO "LINKED_LIST_LENGTH" DO
       IF #list.me[#pointer_list].meta.key = "NULL_TOKEN" THEN
           #ret := INT_TO_DINT(#pointer_list);
           EXIT;
       END_IF;
   END_FOR;
   #"Linked List: Private: Next Empty Node" := #ret;
END_FUNCTION

FUNCTION "Linked List: Append" : Void   // FC169, SCL
{ S7_Optimized_Access := 'TRUE' }
VERSION : 0.1
   VAR_INPUT
      terminal_behavior : String;
   END_VAR
   VAR_IN_OUT
      commands : "Linked List: Method Interface: Append";
      list : "Linked List: List";
   END_VAR
   VAR_TEMP
      clear_commands : "Linked List: Method Interface: Append";
      head : "Linked List: Node";
      pointer_new_node : DInt;
      tail : "Linked List: Node";
   END_VAR
   VAR CONSTANT
      no_error : String := 'no error';
      list_full : String := 'appended to full list';
      no_tail_found : String := 'no tail found while trying to append';
      appended_as_head : String := 'appended as head of list';
   END_VAR
BEGIN
   REGION "NOTES"
       (*
       Append adds a node to the end of the list.
       Last edit: 2021-10-05
       *)
   END_REGION

   REGION "APPEND TO FULL LIST"
       IF "Linked List: Private: Is Full"(#list) THEN
           #commands := #clear_commands;
           #commands.out.error := TRUE;
           #commands.out.error_message := #list_full;
           RETURN;
       END_IF;
   END_REGION

   REGION "APPEND TO EMPTY LIST"
       IF "Linked List: Private: Is Empty"(#list) THEN
           "Linked List: Private: Head an Empty List"(data := #commands.in.data,
                                                      terminal_behavior := #terminal_behavior,
                                                      list := #list);
           #commands := #clear_commands;
           #commands.out.done := TRUE;
           #commands.out.error_message := #appended_as_head;
           RETURN;
       END_IF;
   END_REGION

   REGION "FIND TAIL"
       #tail := "Linked List: Private: Get Tail"(#list);
   END_REGION

   REGION "EXIT CONDITION: TAIL NOT FOUND"
       IF #tail.meta.key = "NULL_TOKEN" THEN
           #commands := #clear_commands;
           #commands.out.error := TRUE;
           #commands.out.error_message := #no_tail_found;
           RETURN;
       END_IF;
   END_REGION

   REGION "FIND FIRST NULL"
       #pointer_new_node := "Linked List: Private: Next Empty Node"(#list);
   END_REGION

   REGION "APPENDED NODE IS AFTER TAIL"
       #list.me[#pointer_new_node].data := #commands.in.data;
       #list.me[#pointer_new_node].meta.key := #pointer_new_node;
       "Linked List: Private: After"(node := #list.me[#pointer_new_node],
                                     previous_node := #list.me[#tail.meta.key]);
   END_REGION

   REGION "EXIT CONDITION: SUCCESS"
       #commands := #clear_commands;
       #commands.out.done := TRUE;
       #commands.out.error_message := #no_error;
   END_REGION
END_FUNCTION

FUNCTION "Linked List: Delete" : Void   // FC170, SCL
{ S7_Optimized_Access := 'TRUE' }
VERSION : 0.1
   VAR_IN_OUT
      commands : "Linked List: Method Interface: Delete";
      list : "Linked List: List";
   END_VAR
   VAR_TEMP
      blank_node : "Linked List: Node";
      clear_commands : "Linked List: Method Interface: Delete";
      current : "Linked List: Node";
      found : Bool;
      next : "Linked List: Node";
      pointer_list : DInt;
      previous : "Linked List: Node";
      search_commands : "Linked List: Method Interface: Search";
   END_VAR
   VAR CONSTANT
      no_error : String := 'no error';
      delete_from_empty : String := 'deleted from an empty list.';
   END_VAR
BEGIN
   REGION "EXIT CONDITION: LIST IS EMPTY"
       IF "Linked List: Private: Is Empty"(#list) THEN
           #commands := #clear_commands;
           #commands.out.error := TRUE;
           #commands.out.error_message := #delete_from_empty;
       END_IF;
   END_REGION

   REGION "DELETE"
       #current := #commands.in.node;
       #previous := "Linked List: Private: Get Previous"(current := #current,
                                                         list := #list);
       #next := "Linked List: Private: Get Next"(current := #current,
                                                 list := #list);
       IF #current.meta.is_head AND NOT #current.meta.is_tail THEN
           "Linked List: Private: Head Swap"(new_head := #list.me[#next.meta.key],
                                             old_head := #list.me[#current.meta.key]);
       END_IF;
       IF NOT #current.meta.is_head AND #current.meta.is_tail THEN
           "Linked List: Private: Tail Swap"(new_tail := #list.me[#previous.meta.key],
                                             old_tail := #list.me[#current.meta.key]);
       END_IF;
       IF NOT #current.meta.is_head THEN
           #list.me[#previous.meta.key].meta.next := #next.meta.key;
       END_IF;
       "Linked List: Private: Clear Node"(#list.me[#current.meta.key]);
   END_REGION

   REGION "COMMANDS OUT"
       #commands := #clear_commands;
       #commands.out.done := TRUE;
       #commands.out.error_message := #no_error;
   END_REGION
END_FUNCTION

FUNCTION "Linked List: Search" : Void   // FC171, SCL
{ S7_Optimized_Access := 'TRUE' }
VERSION : 0.1
   VAR_IN_OUT
      commands : "Linked List: Method Interface: Search";
      list : "Linked List: List";
   END_VAR
   VAR_TEMP
      clear_commands : "Linked List: Method Interface: Search";
      found : Bool;
      pointer_list : DInt;
   END_VAR
   VAR CONSTANT
      no_error : String := 'no error';
      searched_empty_list : String := 'searched empty list';
   END_VAR
BEGIN
   REGION "EXIT CONDITION: SEARCHED EMPTY LIST"
       IF "Linked List: Private: Is Empty"(#list) THEN
           #commands := #clear_commands;
           #commands.out.not_found := TRUE;
           #commands.out.error := TRUE;
           #commands.out.error_message := #searched_empty_list;
           RETURN;
       END_IF;
   END_REGION

   REGION "SEARCH"
       FOR #pointer_list := 0 TO "LINKED_LIST_LENGTH" DO
           IF #list.me[#pointer_list].data = #commands.in.data THEN
               #found := TRUE;
               EXIT;
           END_IF;
       END_FOR;
   END_REGION

   REGION "FOUND"
       IF #found THEN
           #commands := #clear_commands;
           #commands.out.done := TRUE;
           #commands.out.found := TRUE;
           #commands.out.returned_node := #list.me[#pointer_list];
           #commands.out.error_message := #no_error;
           RETURN;
       END_IF;
   END_REGION

   REGION "NOT FOUND"
       IF NOT #found THEN
           #commands := #clear_commands;
           #commands.out.done := TRUE;
           #commands.out.not_found := TRUE;
           RETURN;
       END_IF;
   END_REGION
END_FUNCTION

FUNCTION "Linked List: Display" : Void   // FC172, SCL
{ S7_Optimized_Access := 'TRUE' }
VERSION : 0.1
   VAR_IN_OUT
      commands : "Linked List: Method Interface: Display";
      list : "Linked List: List";
   END_VAR
   VAR_TEMP
      clear_commands : "Linked List: Method Interface: Display";
   END_VAR
BEGIN
   #commands := #clear_commands;
   #commands.out.list := #list;
   #commands.out.done := TRUE;
END_FUNCTION

FUNCTION "Linked List: Insert" : Void   // FC173, SCL
{ S7_Optimized_Access := 'TRUE' }
VERSION : 0.1
   VAR_INPUT
      terminal_behavior : String;
   END_VAR
   VAR_IN_OUT
      commands : "Linked List: Method Interface: Insert";
      list : "Linked List: List";
   END_VAR
   VAR_TEMP
      clear_commands : "Linked List: Method Interface: Insert";
      current : "Linked List: Node";
      next_empty_node_index : DInt;
      previous : "Linked List: Node";
      next : "Linked List: Node";
   END_VAR
   VAR CONSTANT
      no_error : String := 'no error';
      inserted_into_full : String := 'attempted to insert into full list. delete a node and try again.';
      appended_as_head : String := 'appended as head of list';
   END_VAR
BEGIN
   REGION "EXIT CONDITION: INSERTED INTO FULL LIST"
       IF "Linked List: Private: Is Full"(#list) THEN
           #commands := #clear_commands;
           #commands.out.error := TRUE;
           #commands.out.error_message := #inserted_into_full;
           RETURN;
       END_IF;
   END_REGION

   REGION "EXIT CONDITION: INSERTED INTO EMPTY LIST"
       IF "Linked List: Private: Is Empty"(#list) THEN
           "Linked List: Private: Head an Empty List"(data := #commands.in.data,
                                                      terminal_behavior := #terminal_behavior,
                                                      list := #list);
           #commands := #clear_commands;
           #commands.out.error := TRUE;
           #commands.out.error_message := #appended_as_head;
           RETURN;
       END_IF;
   END_REGION

   REGION "GET INDEX OF NEXT EMPTY NODE"
       #next_empty_node_index := "Linked List: Private: Next Empty Node"(#list);
   END_REGION

   REGION "PREVIOUS, CURRENT, AND NEXT NODES"
       #current := #commands.in.target_node;
       #previous := "Linked List: Private: Get Previous"(current := #current,
                                                         list := #list);
       #next := #current;
   END_REGION

   REGION "INSERT BEFORE TARGET NODE"
       // new node's data becomes command data
       #list.me[#next_empty_node_index].data := #commands.in.data;
       // new node's key becomes array index
       #list.me[#next_empty_node_index].meta.key := #next_empty_node_index;
       // shorten name for indexing
       #current := #list.me[#next_empty_node_index];
       // insert
       IF NOT #next.meta.is_head THEN
           "Linked List: Private: After"(node := #list.me[#current.meta.key],
                                         previous_node := #list.me[#previous.meta.key]);
       END_IF;
       "Linked List: Private: Before"(next_node := #list.me[#next.meta.key],
                                      node := #list.me[#current.meta.key]);
   END_REGION

   REGION "COMMANDS OUT"
       #commands := #clear_commands;
       #commands.out.done := TRUE;
       #commands.out.error_message := #no_error;
   END_REGION
END_FUNCTION

FUNCTION "Linked List: Reverse" : Void   // FC174, SCL
{ S7_Optimized_Access := 'TRUE' }